   "Carrier_19_G120DStatusWord.6" AT %I1312.6 : Bool;   // Bit_06_LOCK_OUT
   "Carrier_19_G120DStatusWord.7" AT %I1312.7 : Bool;   // Bit_07_WARN
   "Carrier_19_G120DStatusWord.8" AT %I1313.0 : Bool;   // Bit_08_NO_DEVIATION
   "Carrier_19_G120DStatusWord.9" AT %I1313.1 : Bool;   // Bit_09_CONTR_PLC
   "Carrier_19_G120DStatusWord.10" AT %I1313.2 : Bool;   // Bit_10_F_MAX
   "Carrier_19_G120DStatusWord.11" AT %I1313.3 : Bool;   // Bit_11_LIMIT_REACHED
   "Carrier_19_G120DStatusWord.12" AT %I1313.4 : Bool;   // Bit_12_BRAKE_OPEN
   "Carrier_19_G120DStatusWord.13" AT %I1313.5 : Bool;   // Bit_13_NO_OVERTEMP
   "Carrier_19_G120DStatusWord.14" AT %I1313.6 : Bool;   // Bit_14_CW_CCW
   "Carrier_19_G120DStatusWord.15" AT %I1313.7 : Bool;   // Bit_15_OVERL
   "Carrier_19_Slot2_Input" AT %IW1314 : Word;   // SLOT 2 INPUT WORD
   "Carrier_19_CrashDetectSW" AT %I1314.0 : Bool;   // CRASH DETECT SW
   "Carrier_19_SpareSafetyInput(2_1)" AT %I1314.1 : Bool;   // SPARE SAFETY INPUT
   "Carrier_19_SpareSafetyInput(2_2)" AT %I1314.2 : Bool;   // SPARE SAFETY INPUT
   "Carrier_19_SpareSafetyInput(2_3)" AT %I1314.3 : Bool;   // SPARE SAFETY INPUT
   "Carrier_19_SpareSafetyInput(2_4)" AT %I1314.4 : Bool;   // SPARE SAFETY INPUT
   "Carrier_19_SpareSafetyInput(2_5)" AT %I1314.5 : Bool;   // SPARE SAFETY INPUT
   "Carrier_19_SpareSafetyInput(2_6)" AT %I1314.6 : Bool;   // SPARE SAFETY INPUT
   "Carrier_19_SpareSafetyInput(2_7)" AT %I1314.7 : Bool;   // SPARE SAFETY INPUT
   "Carrier_19_Slot3_SafetyOutput" AT %IW1315 : Word;   // SLOT 3 SAFETY OUTPUT WORD
   "Carrier_19_Crash_Detect_OK" AT %I1315.0 : Bool;   // CARRIER CRASH DETECT
   "Carrier_19_SpareSafetyOutput(3_1)" AT %I1315.1 : Bool;   // SPARE SAFETY OUTPUT
   "Carrier_19_SpareSafetyOutput(3_2)" AT %I1315.2 : Bool;   // SPARE SAFETY OUTPUT
   "Carrier_19_SpareSafetyOutput(3_3)" AT %I1315.3 : Bool;   // SPARE SAFETY OUTPUT
   "Carrier_19_SpareSafetyOutput(3_4)" AT %I1315.4 : Bool;   // SPARE SAFETY OUTPUT
   "Carrier_19_SpareSafetyOutput(3_5)" AT %I1315.5 : Bool;   // SPARE SAFETY OUTPUT
   "Carrier_19_SpareSafetyOutput(3_6)" AT %I1315.6 : Bool;   // SPARE SAFETY OUTPUT
   "Carrier_19_SpareSafetyOutput(3_7)" AT %I1315.7 : Bool;   // SPARE SAFETY OUTPUT
   "Carrier_19_Slot4_Input" AT %IW1316 : Word;   // SLOT 4 INPUT WORD
   "Carrier_19_480VPowerOn_MDCB1" AT %I1316.0 : Bool;   // 480 VAC POWER ON MDCB 1
   "Carrier_19_SpareInput(4_1)" AT %I1316.1 : Bool;   // SPARE INPUT
   "Carrier_19_SpareInput(4_2)" AT %I1316.2 : Bool;   // SPARE INPUT
   "Carrier_19_SitopSelectStatus" AT %I1316.3 : Bool;   // SITOP SELECT STATUS
   "Carrier_19_DCsupplyOnPSCB2" AT %I1316.4 : Bool;   // DC SUPPLY ON PSCB 2
   "Carrier_19_SpareInput(4_5)" AT %I1316.5 : Bool;   // SPARE INPUT
   "Carrier_19_SpareInput(4_6)" AT %I1316.6 : Bool;   // SPARE INPUT
   "Carrier_19_SpareInput(4_7)" AT %I1316.7 : Bool;   // SPARE INPUT
   "Carrier_19_PB1_ProdHoldLH" AT %I1317.0 : Bool;   // PB 1 PRODUCTION HOLD LH
   "Carrier_19_PB2_ResetLH" AT %I1317.1 : Bool;   // PB 2 RESET LH
   "Carrier_19_PB3_ProdHoldRH" AT %I1317.2 : Bool;   // PB 3 PRODUCTION HOLD RH
   "Carrier_19_PB4_ResetRH" AT %I1317.3 : Bool;   // PB 4 RESET RH
   "Carrier_19_SpareInput(4_14)" AT %I1317.4 : Bool;   // SPARE INPUT
   "Carrier_19_SpareInput(4_15)" AT %I1317.5 : Bool;   // SPARE INPUT
   "Carrier_19_SpareInput(4_16)" AT %I1317.6 : Bool;   // SPARE INPUT
   "Carrier_19_SpareInput(4_17)" AT %I1317.7 : Bool;   // SPARE INPUT
   "Carrier_19_Slot5_Output" AT %IW1318 : Word;   // SLOT 5 OUTPUT WORD
   "Carrier_19_IRD400_HMI_24VDC_ENABLE" AT %I1318.0 : Bool;   // IRD 400 PANEL HMI 24V DC POWER
   "Carrier_19_FaultLight_LH" AT %I1318.1 : Bool;   // FAULT LIGHT LH
   "Carrier_19_RunLight_LH" AT %I1318.2 : Bool;   // RUN LIGHT LH
   "Carrier_19_FaultLight_RH" AT %I1318.3 : Bool;   // FAULT LIGHT RH
   "Carrier_19_RunLight_RH" AT %I1318.4 : Bool;   // RUN LIGHT RH
   "Carrier_19_SpareOutput(5_5)" AT %I1318.5 : Bool;   // SPARE OUTPUT
   "Carrier_19_SpareOutput(5_6)" AT %I1318.6 : Bool;   // SPARE OUTPUT
   "Carrier_19_SpareOutput(5_7)" AT %I1318.7 : Bool;   // SPARE OUTPUT
   "Carrier_19_ActualSpeed" AT %IW1320 : Word;   // ACTUAL SPEED
   "Carrier_19_CarrierDriveAlarm" AT %IW1322 : Word;   // CARRIER DRIVE ALARM
   "Carrier_19_CarrierDriveWarning" AT %IW1324 : Word;   // CARRIER DRIVE WARNING
   "Carrier_20_Status" AT %IW1350 : Word;   // CARRIER STATUS WORD
   "Carrier_20_Status.0" AT %I1350.0 : Bool;   // HEARTBEAT
   "Carrier_20_Status.1" AT %I1350.1 : Bool;   // MANUAL
   "Carrier_20_Status.2" AT %I1350.2 : Bool;   // IN_AUTO
   "Carrier_20_Status.3" AT %I1350.3 : Bool;   // POSITIONING_COMPLETE
   "Carrier_20_Status.4" AT %I1350.4 : Bool;   // PRODUCTION HOLD
   "Carrier_20_Status.5" AT %I1350.5 : Bool;   // CARRIER MOVING FORWARD
   "Carrier_20_Status.6" AT %I1350.6 : Bool;   // CARRIER MOVING REVERSE
   "Carrier_20_Status.7" AT %I1350.7 : Bool;   // CARRIER FAULT
   "Carrier_20_Status.8" AT %I1351.0 : Bool;   // CRASH DETECT TRIPPED
   "Carrier_20_Status.9" AT %I1351.1 : Bool;
   "Carrier_20_Status.10" AT %I1351.2 : Bool;
   "Carrier_20_Status.11" AT %I1351.3 : Bool;
   "Carrier_20_Status.12" AT %I1351.4 : Bool;
   "Carrier_20_Status.13" AT %I1351.5 : Bool;
   "Carrier_20_Status.14" AT %I1351.6 : Bool;
   "Carrier_20_Status.15" AT %I1351.7 : Bool;
   "Carrier_20_SDCFaultCode" AT %IW1352 : Word;   // SDC FAULT CODE
   "Carrier_20_CarrierPosition" AT %ID1354 : DWord;   // CARRIER POSITION
   "Carrier_20_CarrierNumber" AT %IW1358 : Word;   // CARRIER NUMBER
   "Carrier_20_G120DControlWord" AT %IW1360 : Word;   // G120D_STW1_CONTROL
   "Carrier_20_G120DControlWord.0" AT %I1360.0 : Bool;   // Bit_00_ON
   "Carrier_20_G120DControlWord.1" AT %I1360.1 : Bool;   // Bit_01_AUS2_INH
   "Carrier_20_G120DControlWord.2" AT %I1360.2 : Bool;   // Bit_02_AUS3_STOP
   "Carrier_20_G120DControlWord.3" AT %I1360.3 : Bool;   // Bit_03_EN
   "Carrier_20_G120DControlWord.4" AT %I1360.4 : Bool;   // Bit_04_EN_RAMP
   "Carrier_20_G120DControlWord.5" AT %I1360.5 : Bool;   // Bit_05_START_RAMP
   "Carrier_20_G120DControlWord.6" AT %I1360.6 : Bool;   // Bit_06_SETPOINT
   "Carrier_20_G120DControlWord.7" AT %I1360.7 : Bool;   // Bit_07_RESET
   "Carrier_20_G120DControlWord.8" AT %I1361.0 : Bool;   // Bit_08_JOG_R
   "Carrier_20_G120DControlWord.9" AT %I1361.1 : Bool;   // Bit_09_JOG_L
   "Carrier_20_G120DControlWord.10" AT %I1361.2 : Bool;   // Bit_10_CONTR_PLC
   "Carrier_20_G120DControlWord.11" AT %I1361.3 : Bool;   // Bit_11_REVERSE
   "Carrier_20_G120DControlWord.12" AT %I1361.4 : Bool;   // Bit_12_BRAKE_RELEASE
   "Carrier_20_G120DControlWord.13" AT %I1361.5 : Bool;   // Bit_13_DDS
   "Carrier_20_G120DControlWord.14" AT %I1361.6 : Bool;   // Bit_14_DO0
   "Carrier_20_G120DControlWord.15" AT %I1361.7 : Bool;   // Bit_15_DO1
   "Carrier_20_G120DStatusWord" AT %IW1362 : Word;   // G120D_ZSW1_STATUS
   "Carrier_20_G120DStatusWord.0" AT %I1362.0 : Bool;   // Bit_00_READY_RUN
   "Carrier_20_G120DStatusWord.1" AT %I1362.1 : Bool;   // Bit_01_READY_ON
   "Carrier_20_G120DStatusWord.2" AT %I1362.2 : Bool;   // Bit_02_ENABLE
   "Carrier_20_G120DStatusWord.3" AT %I1362.3 : Bool;   // Bit_03_FAULT
   "Carrier_20_G120DStatusWord.4" AT %I1362.4 : Bool;   // Bit_04_OFF2
   "Carrier_20_G120DStatusWord.5" AT %I1362.5 : Bool;   // Bit_05_OFF3
   "Carrier_20_G120DStatusWord.6" AT %I1362.6 : Bool;   // Bit_06_LOCK_OUT
   "Carrier_20_G120DStatusWord.7" AT %I1362.7 : Bool;   // Bit_07_WARN
   "Carrier_20_G120DStatusWord.8" AT %I1363.0 : Bool;   // Bit_08_NO_DEVIATION
   "Carrier_20_G120DStatusWord.9" AT %I1363.1 : Bool;   // Bit_09_CONTR_PLC
   "Carrier_20_G120DStatusWord.10" AT %I1363.2 : Bool;   // Bit_10_F_MAX
   "Carrier_20_G120DStatusWord.11" AT %I1363.3 : Bool;   // Bit_11_LIMIT_REACHED
   "Carrier_20_G120DStatusWord.12" AT %I1363.4 : Bool;   // Bit_12_BRAKE_OPEN
   "Carrier_20_G120DStatusWord.13" AT %I1363.5 : Bool;   // Bit_13_NO_OVERTEMP
   "Carrier_20_G120DStatusWord.14" AT %I1363.6 : Bool;   // Bit_14_CW_CCW
   "Carrier_20_G120DStatusWord.15" AT %I1363.7 : Bool;   // Bit_15_OVERL
   "Carrier_20_Slot2_Input" AT %IW1364 : Word;   // SLOT 2 INPUT WORD
   "Carrier_20_CrashDetectSW" AT %I1364.0 : Bool;   // CRASH DETECT SW
   "Carrier_20_SpareSafetyInput(2_1)" AT %I1364.1 : Bool;   // SPARE SAFETY INPUT
   "Carrier_20_SpareSafetyInput(2_2)" AT %I1364.2 : Bool;   // SPARE SAFETY INPUT
   "Carrier_20_SpareSafetyInput(2_3)" AT %I1364.3 : Bool;   // SPARE SAFETY INPUT
   "Carrier_20_SpareSafetyInput(2_4)" AT %I1364.4 : Bool;   // SPARE SAFETY INPUT
   "Carrier_20_SpareSafetyInput(2_5)" AT %I1364.5 : Bool;   // SPARE SAFETY INPUT
   "Carrier_20_SpareSafetyInput(2_6)" AT %I1364.6 : Bool;   // SPARE SAFETY INPUT
   "Carrier_20_SpareSafetyInput(2_7)" AT %I1364.7 : Bool;   // SPARE SAFETY INPUT
   "Carrier_20_Slot3_SafetyOutput" AT %IW1365 : Word;   // SLOT 3 SAFETY OUTPUT WORD
   "Carrier_20_Crash_Detect_OK" AT %I1365.0 : Bool;   // CARRIER CRASH DETECT
   "Carrier_20_SpareSafetyOutput(3_1)" AT %I1365.1 : Bool;   // SPARE SAFETY OUTPUT
   "Carrier_20_SpareSafetyOutput(3_2)" AT %I1365.2 : Bool;   // SPARE SAFETY OUTPUT
   "Carrier_20_SpareSafetyOutput(3_3)" AT %I1365.3 : Bool;   // SPARE SAFETY OUTPUT
   "Carrier_20_SpareSafetyOutput(3_4)" AT %I1365.4 : Bool;   // SPARE SAFETY OUTPUT
   "Carrier_20_SpareSafetyOutput(3_5)" AT %I1365.5 : Bool;   // SPARE SAFETY OUTPUT
   "Carrier_20_SpareSafetyOutput(3_6)" AT %I1365.6 : Bool;   // SPARE SAFETY OUTPUT
   "Carrier_20_SpareSafetyOutput(3_7)" AT %I1365.7 : Bool;   // SPARE SAFETY OUTPUT
   "Carrier_20_Slot4_Input" AT %IW1366 : Word;   // SLOT 4 INPUT WORD
   "Carrier_20_480VPowerOn_MDCB1" AT %I1366.0 : Bool;   // 480 VAC POWER ON MDCB 1
   "Carrier_20_SpareInput(4_1)" AT %I1366.1 : Bool;   // SPARE INPUT
   "Carrier_20_SpareInput(4_2)" AT %I1366.2 : Bool;   // SPARE INPUT
   "Carrier_20_SitopSelectStatus" AT %I1366.3 : Bool;   // SITOP SELECT STATUS
   "Carrier_20_DCsupplyOnPSCB2" AT %I1366.4 : Bool;   // DC SUPPLY ON PSCB 2
   "Carrier_20_SpareInput(4_5)" AT %I1366.5 : Bool;   // SPARE INPUT
   "Carrier_20_SpareInput(4_6)" AT %I1366.6 : Bool;   // SPARE INPUT
   "Carrier_20_SpareInput(4_7)" AT %I1366.7 : Bool;   // SPARE INPUT
   "Carrier_20_PB1_ProdHoldLH" AT %I1367.0 : Bool;   // PB 1 PRODUCTION HOLD LH
   "Carrier_20_PB2_ResetLH" AT %I1367.1 : Bool;   // PB 2 RESET LH
   "Carrier_20_PB3_ProdHoldRH" AT %I1367.2 : Bool;   // PB 3 PRODUCTION HOLD RH
   "Carrier_20_PB4_ResetRH" AT %I1367.3 : Bool;   // PB 4 RESET RH
   "Carrier_20_SpareInput(4_14)" AT %I1367.4 : Bool;   // SPARE INPUT
   "Carrier_20_SpareInput(4_15)" AT %I1367.5 : Bool;   // SPARE INPUT
   "Carrier_20_SpareInput(4_16)" AT %I1367.6 : Bool;   // SPARE INPUT
   "Carrier_20_SpareInput(4_17)" AT %I1367.7 : Bool;   // SPARE INPUT
   "Carrier_20_Slot5_Output" AT %IW1368 : Word;   // SLOT 5 OUTPUT WORD
   "Carrier_20_IRD400_HMI_24VDC_ENABLE" AT %I1368.0 : Bool;   // IRD 400 PANEL HMI 24V DC POWER
   "Carrier_20_FaultLight_LH" AT %I1368.1 : Bool;   // FAULT LIGHT LH
   "Carrier_20_RunLight_LH" AT %I1368.2 : Bool;   // RUN LIGHT LH
   "Carrier_20_FaultLight_RH" AT %I1368.3 : Bool;   // FAULT LIGHT RH
   "Carrier_20_RunLight_RH" AT %I1368.4 : Bool;   // RUN LIGHT RH
   "Carrier_20_SpareOutput(5_5)" AT %I1368.5 : Bool;   // SPARE OUTPUT
   "Carrier_20_SpareOutput(5_6)" AT %I1368.6 : Bool;   // SPARE OUTPUT
   "Carrier_20_SpareOutput(5_7)" AT %I1368.7 : Bool;   // SPARE OUTPUT
   "Carrier_20_ActualSpeed" AT %IW1370 : Word;   // ACTUAL SPEED
   "Carrier_20_CarrierDriveAlarm" AT %IW1372 : Word;   // CARRIER DRIVE ALARM
   "Carrier_20_CarrierDriveWarning" AT %IW1374 : Word;   // CARRIER DRIVE WARNING
   "Carrier_21_Status" AT %IW1400 : Word;   // CARRIER STATUS WORD
   "Carrier_21_Status.0" AT %I1400.0 : Bool;   // HEARTBEAT
   "Carrier_21_Status.1" AT %I1400.1 : Bool;   // MANUAL
   "Carrier_21_Status.2" AT %I1400.2 : Bool;   // IN_AUTO
   "Carrier_21_Status.3" AT %I1400.3 : Bool;   // POSITIONING_COMPLETE
   "Carrier_21_Status.4" AT %I1400.4 : Bool;   // PRODUCTION HOLD
   "Carrier_21_Status.5" AT %I1400.5 : Bool;   // CARRIER MOVING FORWARD
   "Carrier_21_Status.6" AT %I1400.6 : Bool;   // CARRIER MOVING REVERSE
   "Carrier_21_Status.7" AT %I1400.7 : Bool;   // CARRIER FAULT
   "Carrier_21_Status.8" AT %I1401.0 : Bool;   // CRASH DETECT TRIPPED
   "Carrier_21_Status.9" AT %I1401.1 : Bool;
   "Carrier_21_Status.10" AT %I1401.2 : Bool;
   "Carrier_21_Status.11" AT %I1401.3 : Bool;
   "Carrier_21_Status.12" AT %I1401.4 : Bool;
   "Carrier_21_Status.13" AT %I1401.5 : Bool;
   "Carrier_21_Status.14" AT %I1401.6 : Bool;
   "Carrier_21_Status.15" AT %I1401.7 : Bool;
   "Carrier_21_SDCFaultCode" AT %IW1402 : Word;   // SDC FAULT CODE
   "Carrier_21_CarrierPosition" AT %ID1404 : DWord;   // CARRIER POSITION
   "Carrier_21_CarrierNumber" AT %IW1408 : Word;   // CARRIER NUMBER
   "Carrier_21_G120DControlWord" AT %IW1410 : Word;   // G120D_STW1_CONTROL
   "Carrier_21_G120DControlWord.0" AT %I1410.0 : Bool;   // Bit_00_ON
   "Carrier_21_G120DControlWord.1" AT %I1410.1 : Bool;   // Bit_01_AUS2_INH
   "Carrier_21_G120DControlWord.2" AT %I1410.2 : Bool;   // Bit_02_AUS3_STOP
   "Carrier_21_G120DControlWord.3" AT %I1410.3 : Bool;   // Bit_03_EN
   "Carrier_21_G120DControlWord.4" AT %I1410.4 : Bool;   // Bit_04_EN_RAMP
   "Carrier_21_G120DControlWord.5" AT %I1410.5 : Bool;   // Bit_05_START_RAMP
   "Carrier_21_G120DControlWord.6" AT %I1410.6 : Bool;   // Bit_06_SETPOINT
   "Carrier_21_G120DControlWord.7" AT %I1410.7 : Bool;   // Bit_07_RESET
   "Carrier_21_G120DControlWord.8" AT %I1411.0 : Bool;   // Bit_08_JOG_R
   "Carrier_21_G120DControlWord.9" AT %I1411.1 : Bool;   // Bit_09_JOG_L
   "Carrier_21_G120DControlWord.10" AT %I1411.2 : Bool;   // Bit_10_CONTR_PLC
   "Carrier_21_G120DControlWord.11" AT %I1411.3 : Bool;   // Bit_11_REVERSE
   "Carrier_21_G120DControlWord.12" AT %I1411.4 : Bool;   // Bit_12_BRAKE_RELEASE
   "Carrier_21_G120DControlWord.13" AT %I1411.5 : Bool;   // Bit_13_DDS
   "Carrier_21_G120DControlWord.14" AT %I1411.6 : Bool;   // Bit_14_DO0
   "Carrier_21_G120DControlWord.15" AT %I1411.7 : Bool;   // Bit_15_DO1
   "Carrier_21_G120DStatusWord" AT %IW1412 : Word;   // G120D_ZSW1_STATUS
   "Carrier_21_G120DStatusWord.0" AT %I1412.0 : Bool;   // Bit_00_READY_RUN
   "Carrier_21_G120DStatusWord.1" AT %I1412.1 : Bool;   // Bit_01_READY_ON
   "Carrier_21_G120DStatusWord.2" AT %I1412.2 : Bool;   // Bit_02_ENABLE
   "Carrier_21_G120DStatusWord.3" AT %I1412.3 : Bool;   // Bit_03_FAULT
   "Carrier_21_G120DStatusWord.4" AT %I1412.4 : Bool;   // Bit_04_OFF2
   "Carrier_21_G120DStatusWord.5" AT %I1412.5 : Bool;   // Bit_05_OFF3
   "Carrier_21_G120DStatusWord.6" AT %I1412.6 : Bool;   // Bit_06_LOCK_OUT
   "Carrier_21_G120DStatusWord.7" AT %I1412.7 : Bool;   // Bit_07_WARN
   "Carrier_21_G120DStatusWord.8" AT %I1413.0 : Bool;   // Bit_08_NO_DEVIATION
   "Carrier_21_G120DStatusWord.9" AT %I1413.1 : Bool;   // Bit_09_CONTR_PLC
   "Carrier_21_G120DStatusWord.10" AT %I1413.2 : Bool;   // Bit_10_F_MAX
   "Carrier_21_G120DStatusWord.11" AT %I1413.3 : Bool;   // Bit_11_LIMIT_REACHED
   "Carrier_21_G120DStatusWord.12" AT %I1413.4 : Bool;   // Bit_12_BRAKE_OPEN
   "Carrier_21_G120DStatusWord.13" AT %I1413.5 : Bool;   // Bit_13_NO_OVERTEMP
   "Carrier_21_G120DStatusWord.14" AT %I1413.6 : Bool;   // Bit_14_CW_CCW
   "Carrier_21_G120DStatusWord.15" AT %I1413.7 : Bool;   // Bit_15_OVERL
   "Carrier_21_Slot2_Input" AT %IW1414 : Word;   // SLOT 2 INPUT WORD
   "Carrier_21_CrashDetectSW" AT %I1414.0 : Bool;   // CRASH DETECT SW
   "Carrier_21_SpareSafetyInput(2_1)" AT %I1414.1 : Bool;   // SPARE SAFETY INPUT
   "Carrier_21_SpareSafetyInput(2_2)" AT %I1414.2 : Bool;   // SPARE SAFETY INPUT
   "Carrier_21_SpareSafetyInput(2_3)" AT %I1414.3 : Bool;   // SPARE SAFETY INPUT
   "Carrier_21_SpareSafetyInput(2_4)" AT %I1414.4 : Bool;   // SPARE SAFETY INPUT
   "Carrier_21_SpareSafetyInput(2_5)" AT %I1414.5 : Bool;   // SPARE SAFETY INPUT
   "Carrier_21_SpareSafetyInput(2_6)" AT %I1414.6 : Bool;   // SPARE SAFETY INPUT
   "Carrier_21_SpareSafetyInput(2_7)" AT %I1414.7 : Bool;   // SPARE SAFETY INPUT
   "Carrier_21_Slot3_SafetyOutput" AT %IW1415 : Word;   // SLOT 3 SAFETY OUTPUT WORD
   "Carrier_21_Crash_Detect_OK" AT %I1415.0 : Bool;   // CARRIER CRASH DETECT
   "Carrier_21_SpareSafetyOutput(3_1)" AT %I1415.1 : Bool;   // SPARE SAFETY OUTPUT
   "Carrier_21_SpareSafetyOutput(3_2)" AT %I1415.2 : Bool;   // SPARE SAFETY OUTPUT
   "Carrier_21_SpareSafetyOutput(3_3)" AT %I1415.3 : Bool;   // SPARE SAFETY OUTPUT
   "Carrier_21_SpareSafetyOutput(3_4)" AT %I1415.4 : Bool;   // SPARE SAFETY OUTPUT
   "Carrier_21_SpareSafetyOutput(3_5)" AT %I1415.5 : Bool;   // SPARE SAFETY OUTPUT
   "Carrier_21_SpareSafetyOutput(3_6)" AT %I1415.6 : Bool;   // SPARE SAFETY OUTPUT
   "Carrier_21_SpareSafetyOutput(3_7)" AT %I1415.7 : Bool;   // SPARE SAFETY OUTPUT
   "Carrier_21_Slot4_Input" AT %IW1416 : Word;   // SLOT 4 INPUT WORD
   "Carrier_21_480VPowerOn_MDCB1" AT %I1416.0 : Bool;   // 480 VAC POWER ON MDCB 1
   "Carrier_21_SpareInput(4_1)" AT %I1416.1 : Bool;   // SPARE INPUT
   "Carrier_21_SpareInput(4_2)" AT %I1416.2 : Bool;   // SPARE INPUT
   "Carrier_21_SitopSelectStatus" AT %I1416.3 : Bool;   // SITOP SELECT STATUS
   "Carrier_21_DCsupplyOnPSCB2" AT %I1416.4 : Bool;   // DC SUPPLY ON PSCB 2
   "Carrier_21_SpareInput(4_5)" AT %I1416.5 : Bool;   // SPARE INPUT
   "Carrier_21_SpareInput(4_6)" AT %I1416.6 : Bool;   // SPARE INPUT
   "Carrier_21_SpareInput(4_7)" AT %I1416.7 : Bool;   // SPARE INPUT
   "Carrier_21_PB1_ProdHoldLH" AT %I1417.0 : Bool;   // PB 1 PRODUCTION HOLD LH
   "Carrier_21_PB2_ResetLH" AT %I1417.1 : Bool;   // PB 2 RESET LH
   "Carrier_21_PB3_ProdHoldRH" AT %I1417.2 : Bool;   // PB 3 PRODUCTION HOLD RH
   "Carrier_21_PB4_ResetRH" AT %I1417.3 : Bool;   // PB 4 RESET RH
   "Carrier_21_SpareInput(4_14)" AT %I1417.4 : Bool;   // SPARE INPUT
   "Carrier_21_SpareInput(4_15)" AT %I1417.5 : Bool;   // SPARE INPUT
   "Carrier_21_SpareInput(4_16)" AT %I1417.6 : Bool;   // SPARE INPUT
   "Carrier_21_SpareInput(4_17)" AT %I1417.7 : Bool;   // SPARE INPUT
   "Carrier_21_Slot5_Output" AT %IW1418 : Word;   // SLOT 5 OUTPUT WORD
   "Carrier_21_IRD400_HMI_24VDC_ENABLE" AT %I1418.0 : Bool;   // IRD 400 PANEL HMI 24V DC POWER
   "Carrier_21_FaultLight_LH" AT %I1418.1 : Bool;   // FAULT LIGHT LH
   "Carrier_21_RunLight_LH" AT %I1418.2 : Bool;   // RUN LIGHT LH
   "Carrier_21_FaultLight_RH" AT %I1418.3 : Bool;   // FAULT LIGHT RH
   "Carrier_21_RunLight_RH" AT %I1418.4 : Bool;   // RUN LIGHT RH
   "Carrier_21_SpareOutput(5_5)" AT %I1418.5 : Bool;   // SPARE OUTPUT
   "Carrier_21_SpareOutput(5_6)" AT %I1418.6 : Bool;   // SPARE OUTPUT
   "Carrier_21_SpareOutput(5_7)" AT %I1418.7 : Bool;   // SPARE OUTPUT
   "Carrier_21_ActualSpeed" AT %IW1420 : Word;   // ACTUAL SPEED
   "Carrier_21_CarrierDriveAlarm" AT %IW1422 : Word;   // CARRIER DRIVE ALARM
   "Carrier_21_CarrierDriveWarning" AT %IW1424 : Word;   // CARRIER DRIVE WARNING
   "Carrier_22_Status" AT %IW1450 : Word;   // CARRIER STATUS WORD
   "Carrier_22_Status.0" AT %I1450.0 : Bool;   // HEARTBEAT
   "Carrier_22_Status.1" AT %I1450.1 : Bool;   // MANUAL
   "Carrier_22_Status.2" AT %I1450.2 : Bool;   // IN_AUTO
   "Carrier_22_Status.3" AT %I1450.3 : Bool;   // POSITIONING_COMPLETE
   "Carrier_22_Status.4" AT %I1450.4 : Bool;   // PRODUCTION HOLD
   "Carrier_22_Status.5" AT %I1450.5 : Bool;   // CARRIER MOVING FORWARD
   "Carrier_22_Status.6" AT %I1450.6 : Bool;   // CARRIER MOVING REVERSE
   "Carrier_22_Status.7" AT %I1450.7 : Bool;   // CARRIER FAULT
   "Carrier_22_Status.8" AT %I1451.0 : Bool;   // CRASH DETECT TRIPPED
   "Carrier_22_Status.9" AT %I1451.1 : Bool;
   "Carrier_22_Status.10" AT %I1451.2 : Bool;
   "Carrier_22_Status.11" AT %I1451.3 : Bool;
   "Carrier_22_Status.12" AT %I1451.4 : Bool;
   "Carrier_22_Status.13" AT %I1451.5 : Bool;
   "Carrier_22_Status.14" AT %I1451.6 : Bool;
   "Carrier_22_Status.15" AT %I1451.7 : Bool;
   "Carrier_22_SDCFaultCode" AT %IW1452 : Word;   // SDC FAULT CODE
   "Carrier_22_CarrierPosition" AT %ID1454 : DWord;   // CARRIER POSITION
   "Carrier_22_CarrierNumber" AT %IW1458 : Word;   // CARRIER NUMBER
   "Carrier_22_G120DControlWord" AT %IW1460 : Word;   // G120D_STW1_CONTROL
   "Carrier_22_G120DControlWord.0" AT %I1460.0 : Bool;   // Bit_00_ON
   "Carrier_22_G120DControlWord.1" AT %I1460.1 : Bool;   // Bit_01_AUS2_INH
   "Carrier_22_G120DControlWord.2" AT %I1460.2 : Bool;   // Bit_02_AUS3_STOP
   "Carrier_22_G120DControlWord.3" AT %I1460.3 : Bool;   // Bit_03_EN
   "Carrier_22_G120DControlWord.4" AT %I1460.4 : Bool;   // Bit_04_EN_RAMP
   "Carrier_22_G120DControlWord.5" AT %I1460.5 : Bool;   // Bit_05_START_RAMP
   "Carrier_22_G120DControlWord.6" AT %I1460.6 : Bool;   // Bit_06_SETPOINT
   "Carrier_22_G120DControlWord.7" AT %I1460.7 : Bool;   // Bit_07_RESET
   "Carrier_22_G120DControlWord.8" AT %I1461.0 : Bool;   // Bit_08_JOG_R
   "Carrier_22_G120DControlWord.9" AT %I1461.1 : Bool;   // Bit_09_JOG_L
   "Carrier_22_G120DControlWord.10" AT %I1461.2 : Bool;   // Bit_10_CONTR_PLC
   "Carrier_22_G120DControlWord.11" AT %I1461.3 : Bool;   // Bit_11_REVERSE
   "Carrier_22_G120DControlWord.12" AT %I1461.4 : Bool;   // Bit_12_BRAKE_RELEASE
   "Carrier_22_G120DControlWord.13" AT %I1461.5 : Bool;   // Bit_13_DDS
   "Carrier_22_G120DControlWord.14" AT %I1461.6 : Bool;   // Bit_14_DO0
   "Carrier_22_G120DControlWord.15" AT %I1461.7 : Bool;   // Bit_15_DO1
   "Carrier_22_G120DStatusWord" AT %IW1462 : Word;   // G120D_ZSW1_STATUS
   "Carrier_22_G120DStatusWord.0" AT %I1462.0 : Bool;   // Bit_00_READY_RUN
   "Carrier_22_G120DStatusWord.1" AT %I1462.1 : Bool;   // Bit_01_READY_ON
   "Carrier_22_G120DStatusWord.2" AT %I1462.2 : Bool;   // Bit_02_ENABLE
   "Carrier_22_G120DStatusWord.3" AT %I1462.3 : Bool;   // Bit_03_FAULT
   "Carrier_22_G120DStatusWord.4" AT %I1462.4 : Bool;   // Bit_04_OFF2
   "Carrier_22_G120DStatusWord.5" AT %I1462.5 : Bool;   // Bit_05_OFF3
   "Carrier_22_G120DStatusWord.6" AT %I1462.6 : Bool;   // Bit_06_LOCK_OUT
   "Carrier_22_G120DStatusWord.7" AT %I1462.7 : Bool;   // Bit_07_WARN
   "Carrier_22_G120DStatusWord.8" AT %I1463.0 : Bool;   // Bit_08_NO_DEVIATION
   "Carrier_22_G120DStatusWord.9" AT %I1463.1 : Bool;   // Bit_09_CONTR_PLC
   "Carrier_22_G120DStatusWord.10" AT %I1463.2 : Bool;   // Bit_10_F_MAX
   "Carrier_22_G120DStatusWord.11" AT %I1463.3 : Bool;   // Bit_11_LIMIT_REACHED
   "Carrier_22_G120DStatusWord.12" AT %I1463.4 : Bool;   // Bit_12_BRAKE_OPEN
   "Carrier_22_G120DStatusWord.13" AT %I1463.5 : Bool;   // Bit_13_NO_OVERTEMP
   "Carrier_22_G120DStatusWord.14" AT %I1463.6 : Bool;   // Bit_14_CW_CCW
   "Carrier_22_G120DStatusWord.15" AT %I1463.7 : Bool;   // Bit_15_OVERL
   "Carrier_22_Slot2_Input" AT %IW1464 : Word;   // SLOT 2 INPUT WORD
   "Carrier_22_CrashDetectSW" AT %I1464.0 : Bool;   // CRASH DETECT SW
   "Carrier_22_SpareSafetyInput(2_1)" AT %I1464.1 : Bool;   // SPARE SAFETY INPUT
   "Carrier_22_SpareSafetyInput(2_2)" AT %I1464.2 : Bool;   // SPARE SAFETY INPUT
   "Carrier_22_SpareSafetyInput(2_3)" AT %I1464.3 : Bool;   // SPARE SAFETY INPUT
   "Carrier_22_SpareSafetyInput(2_4)" AT %I1464.4 : Bool;   // SPARE SAFETY INPUT
   "Carrier_22_SpareSafetyInput(2_5)" AT %I1464.5 : Bool;   // SPARE SAFETY INPUT
   "Carrier_22_SpareSafetyInput(2_6)" AT %I1464.6 : Bool;   // SPARE SAFETY INPUT
   "Carrier_22_SpareSafetyInput(2_7)" AT %I1464.7 : Bool;   // SPARE SAFETY INPUT
   "Carrier_22_Slot3_SafetyOutput" AT %IW1465 : Word;   // SLOT 3 SAFETY OUTPUT WORD
   "Carrier_22_Crash_Detect_OK" AT %I1465.0 : Bool;   // CARRIER CRASH DETECT
   "Carrier_22_SpareSafetyOutput(3_1)" AT %I1465.1 : Bool;   // SPARE SAFETY OUTPUT
   "Carrier_22_SpareSafetyOutput(3_2)" AT %I1465.2 : Bool;   // SPARE SAFETY OUTPUT
   "Carrier_22_SpareSafetyOutput(3_3)" AT %I1465.3 : Bool;   // SPARE SAFETY OUTPUT
   "Carrier_22_SpareSafetyOutput(3_4)" AT %I1465.4 : Bool;   // SPARE SAFETY OUTPUT
   "Carrier_22_SpareSafetyOutput(3_5)" AT %I1465.5 : Bool;   // SPARE SAFETY OUTPUT
   "Carrier_22_SpareSafetyOutput(3_6)" AT %I1465.6 : Bool;   // SPARE SAFETY OUTPUT
   "Carrier_22_SpareSafetyOutput(3_7)" AT %I1465.7 : Bool;   // SPARE SAFETY OUTPUT
   "Carrier_22_Slot4_Input" AT %IW1466 : Word;   // SLOT 4 INPUT WORD
   "Carrier_22_480VPowerOn_MDCB1" AT %I1466.0 : Bool;   // 480 VAC POWER ON MDCB 1
   "Carrier_22_SpareInput(4_1)" AT %I1466.1 : Bool;   // SPARE INPUT
   "Carrier_22_SpareInput(4_2)" AT %I1466.2 : Bool;   // SPARE INPUT
   "Carrier_22_SitopSelectStatus" AT %I1466.3 : Bool;   // SITOP SELECT STATUS
   "Carrier_22_DCsupplyOnPSCB2" AT %I1466.4 : Bool;   // DC SUPPLY ON PSCB 2
   "Carrier_22_SpareInput(4_5)" AT %I1466.5 : Bool;   // SPARE INPUT
   "Carrier_22_SpareInput(4_6)" AT %I1466.6 : Bool;   // SPARE INPUT
   "Carrier_22_SpareInput(4_7)" AT %I1466.7 : Bool;   // SPARE INPUT
   "Carrier_22_PB1_ProdHoldLH" AT %I1467.0 : Bool;   // PB 1 PRODUCTION HOLD LH
   "Carrier_22_PB2_ResetLH" AT %I1467.1 : Bool;   // PB 2 RESET LH
   "Carrier_22_PB3_ProdHoldRH" AT %I1467.2 : Bool;   // PB 3 PRODUCTION HOLD RH
   "Carrier_22_PB4_ResetRH" AT %I1467.3 : Bool;   // PB 4 RESET RH
   "Carrier_22_SpareInput(4_14)" AT %I1467.4 : Bool;   // SPARE INPUT
   "Carrier_22_SpareInput(4_15)" AT %I1467.5 : Bool;   // SPARE INPUT
   "Carrier_22_SpareInput(4_16)" AT %I1467.6 : Bool;   // SPARE INPUT
   "Carrier_22_SpareInput(4_17)" AT %I1467.7 : Bool;   // SPARE INPUT
   "Carrier_22_Slot5_Output" AT %IW1468 : Word;   // SLOT 5 OUTPUT WORD
   "Carrier_22_IRD400_HMI_24VDC_ENABLE" AT %I1468.0 : Bool;   // IRD 400 PANEL HMI 24V DC POWER
   "Carrier_22_FaultLight_LH" AT %I1468.1 : Bool;   // FAULT LIGHT LH
   "Carrier_22_RunLight_LH" AT %I1468.2 : Bool;   // RUN LIGHT LH
   "Carrier_22_FaultLight_RH" AT %I1468.3 : Bool;   // FAULT LIGHT RH
   "Carrier_22_RunLight_RH" AT %I1468.4 : Bool;   // RUN LIGHT RH
   "Carrier_22_SpareOutput(5_5)" AT %I1468.5 : Bool;   // SPARE OUTPUT
   "Carrier_22_SpareOutput(5_6)" AT %I1468.6 : Bool;   // SPARE OUTPUT
   "Carrier_22_SpareOutput(5_7)" AT %I1468.7 : Bool;   // SPARE OUTPUT
   "Carrier_22_ActualSpeed" AT %IW1470 : Word;   // ACTUAL SPEED
   "Carrier_22_CarrierDriveAlarm" AT %IW1472 : Word;   // CARRIER DRIVE ALARM
   "Carrier_22_CarrierDriveWarning" AT %IW1474 : Word;   // CARRIER DRIVE WARNING
   "Carrier_23_Status" AT %IW1500 : Word;   // CARRIER STATUS WORD
   "Carrier_23_Status.0" AT %I1500.0 : Bool;   // HEARTBEAT
   "Carrier_23_Status.1" AT %I1500.1 : Bool;   // MANUAL
   "Carrier_23_Status.2" AT %I1500.2 : Bool;   // IN_AUTO
   "Carrier_23_Status.3" AT %I1500.3 : Bool;   // POSITIONING_COMPLETE
   "Carrier_23_Status.4" AT %I1500.4 : Bool;   // PRODUCTION HOLD
   "Carrier_23_Status.5" AT %I1500.5 : Bool;   // CARRIER MOVING FORWARD
   "Carrier_23_Status.6" AT %I1500.6 : Bool;   // CARRIER MOVING REVERSE
   "Carrier_23_Status.7" AT %I1500.7 : Bool;   // CARRIER FAULT
   "Carrier_23_Status.8" AT %I1501.0 : Bool;   // CRASH DETECT TRIPPED
   "Carrier_23_Status.9" AT %I1501.1 : Bool;
   "Carrier_23_Status.10" AT %I1501.2 : Bool;
   "Carrier_23_Status.11" AT %I1501.3 : Bool;
   "Carrier_23_Status.12" AT %I1501.4 : Bool;
   "Carrier_23_Status.13" AT %I1501.5 : Bool;
   "Carrier_23_Status.14" AT %I1501.6 : Bool;
   "Carrier_23_Status.15" AT %I1501.7 : Bool;
   "Carrier_23_SDCFaultCode" AT %IW1502 : Word;   // SDC FAULT CODE
   "Carrier_23_CarrierPosition" AT %ID1504 : DWord;   // CARRIER POSITION
   "Carrier_23_CarrierNumber" AT %IW1508 : Word;   // CARRIER NUMBER
   "Carrier_23_G120DControlWord" AT %IW1510 : Word;   // G120D_STW1_CONTROL
   "Carrier_23_G120DControlWord.0" AT %I1510.0 : Bool;   // Bit_00_ON
   "Carrier_23_G120DControlWord.1" AT %I1510.1 : Bool;   // Bit_01_AUS2_INH
   "Carrier_23_G120DControlWord.2" AT %I1510.2 : Bool;   // Bit_02_AUS3_STOP
   "Carrier_23_G120DControlWord.3" AT %I1510.3 : Bool;   // Bit_03_EN
   "Carrier_23_G120DControlWord.4" AT %I1510.4 : Bool;   // Bit_04_EN_RAMP
   "Carrier_23_G120DControlWord.5" AT %I1510.5 : Bool;   // Bit_05_START_RAMP
   "Carrier_23_G120DControlWord.6" AT %I1510.6 : Bool;   // Bit_06_SETPOINT
   "Carrier_23_G120DControlWord.7" AT %I1510.7 : Bool;   // Bit_07_RESET
   "Carrier_23_G120DControlWord.8" AT %I1511.0 : Bool;   // Bit_08_JOG_R
   "Carrier_23_G120DControlWord.9" AT %I1511.1 : Bool;   // Bit_09_JOG_L
   "Carrier_23_G120DControlWord.10" AT %I1511.2 : Bool;   // Bit_10_CONTR_PLC
   "Carrier_23_G120DControlWord.11" AT %I1511.3 : Bool;   // Bit_11_REVERSE
   "Carrier_23_G120DControlWord.12" AT %I1511.4 : Bool;   // Bit_12_BRAKE_RELEASE
   "Carrier_23_G120DControlWord.13" AT %I1511.5 : Bool;   // Bit_13_DDS
   "Carrier_23_G120DControlWord.14" AT %I1511.6 : Bool;   // Bit_14_DO0
   "Carrier_23_G120DControlWord.15" AT %I1511.7 : Bool;   // Bit_15_DO1
   "Carrier_23_G120DStatusWord" AT %IW1512 : Word;   // G120D_ZSW1_STATUS
   "Carrier_23_G120DStatusWord.0" AT %I1512.0 : Bool;   // Bit_00_READY_RUN
   "Carrier_23_G120DStatusWord.1" AT %I1512.1 : Bool;   // Bit_01_READY_ON
   "Carrier_23_G120DStatusWord.2" AT %I1512.2 : Bool;   // Bit_02_ENABLE
   "Carrier_23_G120DStatusWord.3" AT %I1512.3 : Bool;   // Bit_03_FAULT
   "Carrier_23_G120DStatusWord.4" AT %I1512.4 : Bool;   // Bit_04_OFF2
   "Carrier_23_G120DStatusWord.5" AT %I1512.5 : Bool;   // Bit_05_OFF3
   "Carrier_23_G120DStatusWord.6" AT %I1512.6 : Bool;   // Bit_06_LOCK_OUT
   "Carrier_23_G120DStatusWord.7" AT %I1512.7 : Bool;   // Bit_07_WARN
   "Carrier_23_G120DStatusWord.8" AT %I1513.0 : Bool;   // Bit_08_NO_DEVIATION
   "Carrier_23_G120DStatusWord.9" AT %I1513.1 : Bool;   // Bit_09_CONTR_PLC
   "Carrier_23_G120DStatusWord.10" AT %I1513.2 : Bool;   // Bit_10_F_MAX
   "Carrier_23_G120DStatusWord.11" AT %I1513.3 : Bool;   // Bit_11_LIMIT_REACHED
   "Carrier_23_G120DStatusWord.12" AT %I1513.4 : Bool;   // Bit_12_BRAKE_OPEN
   "Carrier_23_G120DStatusWord.13" AT %I1513.5 : Bool;   // Bit_13_NO_OVERTEMP
   "Carrier_23_G120DStatusWord.14" AT %I1513.6 : Bool;   // Bit_14_CW_CCW
   "Carrier_23_G120DStatusWord.15" AT %I1513.7 : Bool;   // Bit_15_OVERL
   "Carrier_23_Slot2_Input" AT %IW1514 : Word;   // SLOT 2 INPUT WORD
   "Carrier_23_CrashDetectSW" AT %I1514.0 : Bool;   // CRASH DETECT SW
   "Carrier_23_SpareSafetyInput(2_1)" AT %I1514.1 : Bool;   // SPARE SAFETY INPUT
   "Carrier_23_SpareSafetyInput(2_2)" AT %I1514.2 : Bool;   // SPARE SAFETY INPUT
   "Carrier_23_SpareSafetyInput(2_3)" AT %I1514.3 : Bool;   // SPARE SAFETY INPUT
   "Carrier_23_SpareSafetyInput(2_4)" AT %I1514.4 : Bool;   // SPARE SAFETY INPUT
   "Carrier_23_SpareSafetyInput(2_5)" AT %I1514.5 : Bool;   // SPARE SAFETY INPUT
   "Carrier_23_SpareSafetyInput(2_6)" AT %I1514.6 : Bool;   // SPARE SAFETY INPUT
   "Carrier_23_SpareSafetyInput(2_7)" AT %I1514.7 : Bool;   // SPARE SAFETY INPUT
   "Carrier_23_Slot3_SafetyOutput" AT %IW1515 : Word;   // SLOT 3 SAFETY OUTPUT WORD
   "Carrier_23_Crash_Detect_OK" AT %I1515.0 : Bool;   // CARRIER CRASH DETECT
   "Carrier_23_SpareSafetyOutput(3_1)" AT %I1515.1 : Bool;   // SPARE SAFETY OUTPUT
   "Carrier_23_SpareSafetyOutput(3_2)" AT %I1515.2 : Bool;   // SPARE SAFETY OUTPUT
   "Carrier_23_SpareSafetyOutput(3_3)" AT %I1515.3 : Bool;   // SPARE SAFETY OUTPUT
   "Carrier_23_SpareSafetyOutput(3_4)" AT %I1515.4 : Bool;   // SPARE SAFETY OUTPUT
   "Carrier_23_SpareSafetyOutput(3_5)" AT %I1515.5 : Bool;   // SPARE SAFETY OUTPUT
   "Carrier_23_SpareSafetyOutput(3_6)" AT %I1515.6 : Bool;   // SPARE SAFETY OUTPUT
   "Carrier_23_SpareSafetyOutput(3_7)" AT %I1515.7 : Bool;   // SPARE SAFETY OUTPUT
   "Carrier_23_Slot4_Input" AT %IW1516 : Word;   // SLOT 4 INPUT WORD
   "Carrier_23_480VPowerOn_MDCB1" AT %I1516.0 : Bool;   // 480 VAC POWER ON MDCB 1
   "Carrier_23_SpareInput(4_1)" AT %I1516.1 : Bool;   // SPARE INPUT
   "Carrier_23_SpareInput(4_2)" AT %I1516.2 : Bool;   // SPARE INPUT
   "Carrier_23_SitopSelectStatus" AT %I1516.3 : Bool;   // SITOP SELECT STATUS
   "Carrier_23_DCsupplyOnPSCB2" AT %I1516.4 : Bool;   // DC SUPPLY ON PSCB 2
   "Carrier_23_SpareInput(4_5)" AT %I1516.5 : Bool;   // SPARE INPUT
   "Carrier_23_SpareInput(4_6)" AT %I1516.6 : Bool;   // SPARE INPUT
   "Carrier_23_SpareInput(4_7)" AT %I1516.7 : Bool;   // SPARE INPUT
   "Carrier_23_PB1_ProdHoldLH" AT %I1517.0 : Bool;   // PB 1 PRODUCTION HOLD LH
   "Carrier_23_PB2_ResetLH" AT %I1517.1 : Bool;   // PB 2 RESET LH
   "Carrier_23_PB3_ProdHoldRH" AT %I1517.2 : Bool;   // PB 3 PRODUCTION HOLD RH
   "Carrier_23_PB4_ResetRH" AT %I1517.3 : Bool;   // PB 4 RESET RH
   "Carrier_23_SpareInput(4_14)" AT %I1517.4 : Bool;   // SPARE INPUT
   "Carrier_23_SpareInput(4_15)" AT %I1517.5 : Bool;   // SPARE INPUT
   "Carrier_23_SpareInput(4_16)" AT %I1517.6 : Bool;   // SPARE INPUT
   "Carrier_23_SpareInput(4_17)" AT %I1517.7 : Bool;   // SPARE INPUT
   "Carrier_23_Slot5_Output" AT %IW1518 : Word;   // SLOT 5 OUTPUT WORD
   "Carrier_23_IRD400_HMI_24VDC_ENABLE" AT %I1518.0 : Bool;   // IRD 400 PANEL HMI 24V DC POWER
   "Carrier_23_FaultLight_LH" AT %I1518.1 : Bool;   // FAULT LIGHT LH
   "Carrier_23_RunLight_LH" AT %I1518.2 : Bool;   // RUN LIGHT LH
   "Carrier_23_FaultLight_RH" AT %I1518.3 : Bool;   // FAULT LIGHT RH
   "Carrier_23_RunLight_RH" AT %I1518.4 : Bool;   // RUN LIGHT RH
   "Carrier_23_SpareOutput(5_5)" AT %I1518.5 : Bool;   // SPARE OUTPUT
   "Carrier_23_SpareOutput(5_6)" AT %I1518.6 : Bool;   // SPARE OUTPUT
   "Carrier_23_SpareOutput(5_7)" AT %I1518.7 : Bool;   // SPARE OUTPUT